     "CP_YZ":
       IF (#compDirection = "LKINCTRL_COMP_LEFT") THEN
         #tempVOrthogonal.x := 0.0;
         #tempVOrthogonal.y := - #tempVTangential.z;
         #tempVOrthogonal.z := #tempVTangential.y;
       ELSE
         #tempVOrthogonal.x := 0.0;
         #tempVOrthogonal.y := #tempVTangential.z;
         #tempVOrthogonal.z := - #tempVTangential.y;
       END_IF;
   END_CASE;
   END_REGION CALCULATION

   #vUnitTangentialPathPlane := #tempVTangential;
   #vUnitOrthogonalPathPlane := #tempVOrthogonal;
   #LKinCtrl_CalcLineTangOrthPathPlane := 0;
END_FUNCTION

FUNCTION "LKinCtrl_CalcCircTangOrthPathPlane" : Word   // FC35056, SCL
TITLE = LKinCtrl_CalcCircTangOrthPathPlane
{ S7_Optimized_Access := 'TRUE' }
AUTHOR : tech.team.motioncontrol@siemens.com
FAMILY : LKinCtrl
VERSION : 1.0
// Calculate orthogonal and tangential vector of a circle point with respect ot the path plane
   VAR_INPUT
      circlePoint : "LKinCtrl_typeCOff3DPoint";   // Circle point
      circleCenterPoint : "LKinCtrl_typeCOff3DPoint";   // Circle center point
      pathPlane : Int;   // Path plane: XZ= 0, YZ=1, XY= 2
      compDirection : Int;   // Tool radius compensation direction: left=1, right = 0
      pathChoice : DInt;   // Circle path choice: positive= 0, negative= 1
   END_VAR
   VAR_OUTPUT
      vUnitTangentialPathPlane : "LKinCtrl_typeCOff3DPoint";   // Output tangential vector - path plane - unit vector
      vUnitOrthogonalPathPlane : "LKinCtrl_typeCOff3DPoint";   // Output othogonal vector - path plane - unit vector
   END_VAR
   VAR_TEMP
      tempDiffVec : "LKinCtrl_typeCOff3DPoint";   // Difference vector
      tempVOrthogonal : "LKinCtrl_typeCOff3DPoint";   // Othogonal vector
      tempVTangential : "LKinCtrl_typeCOff3DPoint";   // Tangential vector
   END_VAR
   // Ret_Val : Return value
   VAR CONSTANT
      ERR_COFF_INVALID_PATH_PLANE : Word := 16#8303;   // Error - invalid path plane
      ERR_COFF_INVALID_PATH_CHOICE_OF_CIRCULAR_CMD : Word := 16#8308;   // Error - invalid circle path choice
      ERR_COFF_INVALID_COMPENSATION_DIRECTION : Word := 16#8304;   // Error - invalid compensation direction
   END_VAR
BEGIN
   //=============================================================================
   // SIEMENS AG
   // (c)Copyright 2019 All Rights Reserved
   //-----------------------------------------------------------------------------
   // Library: - 
   // Tested with: S7-1516T-3 PN
   // Engineering: TIA Portal V15
   // Restrictions: -
   // Requirements: S7-1500/S7-1500T FW 2.5
   // Functionality: Calculate orthogonal and tangential vector of a circle point
   // with respect ot the path plane
   //-----------------------------------------------------------------------------
   // Change log table:
   // Version  Date       Expert in charge Changes applied
   // 01.00.00 2019-02-05 AW               created
   //=============================================================================

   REGION PLAUSIBILITY_CHECK
     // Check path plane
     IF ((#pathPlane >= "CP_XZ") AND (#pathPlane <= "CP_XY"))
     THEN
       // Check compensation direction
       IF ((#compDirection >= "LKINCTRL_COMP_LEFT") AND (#compDirection <= "LKINCTRL_COMP_RIGHT"))
       THEN
         // Check compensation direction
         IF ((#pathChoice >= 0) AND (#pathChoice <= 1))
         THEN
           ;
         ELSE
           #LKinCtrl_CalcCircTangOrthPathPlane := #ERR_COFF_INVALID_PATH_CHOICE_OF_CIRCULAR_CMD; // Invalid compensation direction
           RETURN;
         END_IF;
       ELSE
         #LKinCtrl_CalcCircTangOrthPathPlane := #ERR_COFF_INVALID_COMPENSATION_DIRECTION; // Invalid compensation direction
         RETURN;
       END_IF;
     ELSE
       #LKinCtrl_CalcCircTangOrthPathPlane := #ERR_COFF_INVALID_PATH_PLANE; // Invalid path plane
       RETURN;
     END_IF;
   END_REGION PLAUSIBILITY_CHECK

   REGION CALCULATION



     (*
     IF (#compDirection = "LKINCTRL_COMP_LEFT") THEN
       #tempVOrthogonal := "LKinCtrl_VecSub"(vIn1 := #circlePoint, vIn2 := #circleCenterPoint);
     ELSE
       #tempVOrthogonal := "LKinCtrl_VecSub"(vIn1 := #circleCenterPoint, vIn2 := #circlePoint);
     END_IF;
     *)

     // Take care of path plane
     CASE #pathPlane OF
       "CP_XY":
         // Calc radius vector circle center to start point
         IF (#compDirection = "LKINCTRL_COMP_LEFT") THEN
           IF (#pathChoice = 0) THEN
             #tempVOrthogonal := "LKinCtrl_VecSub"(vIn1 := #circleCenterPoint, vIn2 := #circlePoint);
           ELSE
             #tempVOrthogonal := "LKinCtrl_VecSub"(vIn1 := #circlePoint, vIn2 := #circleCenterPoint);
           END_IF;
         ELSE
           IF (#pathChoice = 0) THEN
             #tempVOrthogonal := "LKinCtrl_VecSub"(vIn1 := #circlePoint, vIn2 := #circleCenterPoint);
           ELSE
             #tempVOrthogonal := "LKinCtrl_VecSub"(vIn1 := #circleCenterPoint, vIn2 := #circlePoint);
           END_IF;
         END_IF;
         #tempVOrthogonal.z := 0.0;

       "CP_XZ":
         // Calc radius vector circle center to start point
         IF (#compDirection = "LKINCTRL_COMP_LEFT") THEN
           IF (#pathChoice = 0) THEN
             #tempVOrthogonal := "LKinCtrl_VecSub"(vIn1 := #circlePoint, vIn2 := #circleCenterPoint);
           ELSE
             #tempVOrthogonal := "LKinCtrl_VecSub"(vIn1 := #circleCenterPoint, vIn2 := #circlePoint);
           END_IF;
         ELSE
           IF (#pathChoice = 0) THEN
             #tempVOrthogonal := "LKinCtrl_VecSub"(vIn1 := #circleCenterPoint, vIn2 := #circlePoint);
           ELSE
             #tempVOrthogonal := "LKinCtrl_VecSub"(vIn1 := #circlePoint, vIn2 := #circleCenterPoint);
           END_IF;
         END_IF;
         #tempVOrthogonal.y := 0.0;

       "CP_YZ":
         // Calc radius vector circle center to start point
         IF (#compDirection = "LKINCTRL_COMP_LEFT") THEN
           IF (#pathChoice = 0) THEN
             #tempVOrthogonal := "LKinCtrl_VecSub"(vIn1 := #circleCenterPoint, vIn2 := #circlePoint);
           ELSE
             #tempVOrthogonal := "LKinCtrl_VecSub"(vIn1 := #circlePoint, vIn2 := #circleCenterPoint);
           END_IF;
         ELSE
           IF (#pathChoice = 0) THEN
             #tempVOrthogonal := "LKinCtrl_VecSub"(vIn1 := #circlePoint, vIn2 := #circleCenterPoint);
           ELSE
             #tempVOrthogonal := "LKinCtrl_VecSub"(vIn1 := #circleCenterPoint, vIn2 := #circlePoint);
           END_IF;
         END_IF;
         #tempVOrthogonal.x := 0.0;
     END_CASE;

     #tempVOrthogonal := "LKinCtrl_VecUnit"(#tempVOrthogonal);

     // Check path plane
     IF (#pathPlane = "CP_XY") THEN
       #tempVTangential.x := - #tempVOrthogonal.y;
       #tempVTangential.y := #tempVOrthogonal.x;
       #tempVTangential.z := 0.0;
     ELSIF (#pathPlane = "CP_XZ") THEN
       #tempVTangential.x := #tempVOrthogonal.z;
       #tempVTangential.y := 0.0;
       #tempVTangential.z := - #tempVOrthogonal.x;
     ELSIF (#pathPlane = "CP_YZ") THEN
       #tempVTangential.x := 0.0;
       #tempVTangential.y := - #tempVOrthogonal.z;
       #tempVTangential.z := #tempVOrthogonal.y;
     END_IF;
   END_REGION CALCULATION

   #vUnitTangentialPathPlane := #tempVTangential;
   #vUnitOrthogonalPathPlane := #tempVOrthogonal;

   #LKinCtrl_CalcCircTangOrthPathPlane := 0; // o.k.
END_FUNCTION

FUNCTION "LKinCtrl_CalcCircCenterByIntermediatePointAndEndPoint" : Word   // FC35057, SCL
TITLE = LKinCtrl_CalcCircCenterByIntermediatePointAndEndPoint
{ S7_Optimized_Access := 'TRUE' }
AUTHOR : tech.team.motioncontrol@siemens.com
FAMILY : LKinCtrl
VERSION : 1.0
// Calculate circle center point with given intermediate point
   VAR_INPUT
      circleStartPoint : "LKinCtrl_typeCOff3DPoint";   // Circle start point
      circleEndPoint : "LKinCtrl_typeCOff3DPoint";   // Circle end point
      circleIntermediatePoint : "LKinCtrl_typeCOff3DPoint";   // Circle intermediate point
      pathPlane : Int;   // Path plane: XZ= 0, YZ=1, XY= 2
   END_VAR
   VAR_OUTPUT
      circleCenterPoint : "LKinCtrl_typeCOff3DPoint";   // Circle center point
   END_VAR
   VAR_TEMP
      tempVecL : "LKinCtrl_typeCOff3DPoint";
      tempVecP1P2 : "LKinCtrl_typeCOff3DPoint";
      tempVecP3P4 : "LKinCtrl_typeCOff3DPoint";
      tempLengthVecP1P2 : LReal;
      tempLengthVecP3P4 : LReal;
      tempUnitVecP1P2 : "LKinCtrl_typeCOff3DPoint";
      tempUnitVecP3P4 : "LKinCtrl_typeCOff3DPoint";
      tempP12 : "LKinCtrl_typeCOff3DPoint";
      tempP34 : "LKinCtrl_typeCOff3DPoint";
      tempP123 : "LKinCtrl_typeCOff3DPoint";
      tempP341 : "LKinCtrl_typeCOff3DPoint";
      tempOrthVecP1P2 : "LKinCtrl_typeCOff3DPoint";
      tempOrthVecP3P4 : "LKinCtrl_typeCOff3DPoint";
      tempRetValue : Word;
      tempPa : "LKinCtrl_typeCOff3DPoint";
      tempPb : "LKinCtrl_typeCOff3DPoint";
      tempMua : LReal;
      tempMub : LReal;
   END_VAR
   // Ret_Val : Return value
   VAR CONSTANT
      ERR_COFF_INVALID_PATH_PLANE : Word := 16#8303;   // Error - invalid path plane
   END_VAR
BEGIN
   //=============================================================================
   // SIEMENS AG
   // (c)Copyright 2019 All Rights Reserved
   //-----------------------------------------------------------------------------
   // Library: - 
   // Tested with: S7-1516T-3 PN
   // Engineering: TIA Portal V15
   // Restrictions: -
   // Requirements: S7-1500/S7-1500T FW 2.5
   // Functionality: Calculate circle center point with given intermediate point
   // and end point
   //-----------------------------------------------------------------------------
   // Change log table:
   // Version  Date       Expert in charge Changes applied
   // 01.00.00 2019-02-05 AW               created
   //=============================================================================


   REGION PLAUSIBILITY_CHECK
   // Check path plane
     IF ((#pathPlane >= "CP_XZ") AND (#pathPlane <= "CP_XY"))
   THEN
     ;
   ELSE
     #LKinCtrl_CalcCircCenterByIntermediatePointAndEndPoint := #ERR_COFF_INVALID_PATH_PLANE; // Invalid path plane
     RETURN;
   END_IF;
   END_REGION PLAUSIBILITY_CHECK

   REGION CALCULATION

     // Intermediate point - start point
     #tempVecP1P2 := "LKinCtrl_VecSub"(vIn1:= #circleIntermediatePoint, vIn2:= #circleStartPoint);
     // Intermediate point - end point
     #tempVecP3P4 := "LKinCtrl_VecSub"(vIn1 := #circleIntermediatePoint, vIn2 := #circleEndPoint);

     // Length of vectors
     #tempLengthVecP1P2 := "LKinCtrl_VecAbs"(#tempVecP1P2);
     #tempLengthVecP3P4 := "LKinCtrl_VecAbs"(#tempVecP3P4);

     // Direction of vectors
     #tempUnitVecP1P2 := "LKinCtrl_VecUnit"(#tempVecP1P2);
     #tempUnitVecP3P4 := "LKinCtrl_VecUnit"(#tempVecP3P4);

     // Perpendicular bisector
     #tempP12 := "LKinCtrl_VecAdd"(vIn1:= #circleStartPoint, vIn2:= "LKinCtrl_VecScale"(vIn:= #tempUnitVecP1P2, factor:= (#tempLengthVecP1P2 / 2.0)));
     #tempP34 := "LKinCtrl_VecAdd"(vIn1:= #circleEndPoint, vIn2:="LKinCtrl_VecScale"(vIn:= #tempUnitVecP3P4, factor:=(#tempLengthVecP3P4 / 2.0)));

     // Rotate vector according to path plane
     // Calc complete shift
     CASE #pathPlane OF
       "CP_XY":
           // Orthogonal end point - intermediate point
           #tempOrthVecP1P2.x := - #tempUnitVecP1P2.y;
           #tempOrthVecP1P2.y := #tempUnitVecP1P2.x;
           #tempOrthVecP1P2.z := 0.0;

           // Orthogonal end point - intermediate point
           #tempOrthVecP3P4.x := #tempUnitVecP3P4.y;
           #tempOrthVecP3P4.y := - #tempUnitVecP3P4.x;
           #tempOrthVecP3P4.z := 0.0;

         "CP_XZ":
           // Orthogonal end point - intermediate point
           #tempOrthVecP1P2.x := #tempUnitVecP1P2.z;
           #tempOrthVecP1P2.y := 0.0;
           #tempOrthVecP1P2.z := - #tempUnitVecP1P2.x;

           // Orthogonal end point - intermediate point
           #tempOrthVecP3P4.x := - #tempUnitVecP3P4.z;
           #tempOrthVecP3P4.y := 0.0;
           #tempOrthVecP3P4.z := #tempUnitVecP3P4.x;

         "CP_YZ":
           // Orthogonal end point - intermediate point
           #tempOrthVecP1P2.x := 0.0;
           #tempOrthVecP1P2.y := - #tempUnitVecP1P2.z;
           #tempOrthVecP1P2.z := #tempUnitVecP1P2.y;

           // Orthogonal end point - intermediate point
           #tempOrthVecP3P4.x := 0.0;
           #tempOrthVecP3P4.y := #tempUnitVecP3P4.z;
           #tempOrthVecP3P4.z := - #tempUnitVecP3P4.y;
     END_CASE;

     #tempOrthVecP1P2 := "LKinCtrl_VecScale"(vIn:= #tempOrthVecP1P2, factor:= #tempLengthVecP1P2);
     #tempOrthVecP3P4 := "LKinCtrl_VecScale"(vIn:= #tempOrthVecP3P4, factor:= #tempLengthVecP3P4);

     #tempP123 := "LKinCtrl_VecAdd"(vIn1:= #tempP12, vIn2:= #tempOrthVecP1P2);
     #tempP341 := "LKinCtrl_VecAdd"(vIn1:= #tempP34, vIn2:= #tempOrthVecP3P4);

     #tempRetValue := "LKinCtrl_CalcLineLineIntersectionPoint"(startPointFirstLine := #tempP12,
                                                      endPointFirstLine := #tempP123,
                                                      startPointSecondLine := #tempP34,
                                                      endPointSecondLine := #tempP341,
                                                      intersectionPointA => #tempPa,
                                                      intersectionPointB => #tempPb,
                                                      muA => #tempMua,
                                                      muB => #tempMub);
     IF (#tempRetValue <> 0) THEN
       #LKinCtrl_CalcCircCenterByIntermediatePointAndEndPoint := #tempRetValue;
       RETURN;
     END_IF;

   END_REGION CALCULATION

   #circleCenterPoint := #tempPa;

   #LKinCtrl_CalcCircCenterByIntermediatePointAndEndPoint := 0; // o.k.
END_FUNCTION

FUNCTION "LKinCtrl_CalcCircPathChoiceByIntermediatePointAndEndPoint" : Word   // FC35058, SCL
TITLE = LKinCtrl_CalcCircPathChoiceByIntermediatePointAndEndPoint
{ S7_Optimized_Access := 'TRUE' }
AUTHOR : tech.team.motioncontrol@siemens.com
FAMILY : LKinCtrl
VERSION : 1.0
// Calculate circle path choice by given circle intermediate point and end point
   VAR_INPUT
      circleStartPoint : "LKinCtrl_typeCOff3DPoint";   // Circle start point
      circleEndPoint : "LKinCtrl_typeCOff3DPoint";   // Circle end point
      circleintermediatePoint : "LKinCtrl_typeCOff3DPoint";   // Circle intermediate point
      pathPlane : Int;   // Path plane: XZ= 0, YZ=1, XY= 2
   END_VAR
   VAR_OUTPUT
      pathChoice : DInt;   // Circle path choice: positive= 0, negative= 1
   END_VAR
   VAR_TEMP
      tempVEndStart : "LKinCtrl_typeCOff3DPoint";
      tempVIntStart : "LKinCtrl_typeCOff3DPoint";
      tempCrossVec : "LKinCtrl_typeCOff3DPoint";
   END_VAR
   // Ret_Val : Return value
   VAR CONSTANT
      ERR_COFF_INVALID_PATH_PLANE : Word := 16#8303;   // Error - invalid path plane
   END_VAR
BEGIN
   //=============================================================================
   // SIEMENS AG
   // (c)Copyright 2019 All Rights Reserved
   //-----------------------------------------------------------------------------
   // Library: - 
   // Tested with: S7-1516T-3 PN
   // Engineering: TIA Portal V15
   // Restrictions: -
   // Requirements: S7-1500/S7-1500T FW 2.5
   // Functionality: Calculate circle path choice by given circle intermediate point
   // and end point
   //-----------------------------------------------------------------------------
   // Change log table:
   // Version  Date       Expert in charge Changes applied
   // 01.00.00 2019-02-05 AW               created
   //=============================================================================

   REGION PLAUSIBILITY_CHECK
     // Check path plane
     IF ((#pathPlane >= "CP_XZ") AND (#pathPlane <= "CP_XY"))
     THEN
       ;
     ELSE
       #LKinCtrl_CalcCircPathChoiceByIntermediatePointAndEndPoint := #ERR_COFF_INVALID_PATH_PLANE; // Invalid path plane
       RETURN;
     END_IF;
   END_REGION PLAUSIBILITY_CHECK

   REGION CALCULATION

   (*  
   // Calculate angle between start / end point and start / intermediate point
     #tempRetValue := "LKinCOff_CalcAngleBetweenVectors"(point1 := #endPoint,
                                                         point2 := #intermediatePoint,
                                                         intersectionPoint := #startPoint,
                                                         angle => #tempAngle);


   IF (#tempRetValue <> 0) THEN
     #LKinCOff_CalcPathChoiceByIntermediatePointAndEndPoint := #tempRetValue;
     RETURN;
   END_IF;

   END_REGION CALCULATION
   IF (#tempAngle < 0.0) THEN
     #pathChoice := 1;
   ELSE
     #pathChoice := 0;
   END_IF;
   *)

     // Difference vectors
     #tempVEndStart := "LKinCtrl_VecSub"(vIn1 := #circleEndPoint, vIn2 := #circleStartPoint);
     #tempVIntStart := "LKinCtrl_VecSub"(vIn1 := #circleintermediatePoint, vIn2 := #circleStartPoint);

     #tempCrossVec := "LKinCtrl_VecCrossProd"(vIn1 := #tempVEndStart,
                                              vIn2 := #tempVIntStart);

     // Check path plane
     IF (#pathPlane = "CP_XY") THEN
       IF (#tempCrossVec.z > 0.0) THEN
         #pathChoice := "PC_NEGATIVE";
       ELSE
         #pathChoice := "PC_POSITIVE";
       END_IF;
     ELSIF (#pathPlane = "CP_XZ") THEN
       IF (#tempCrossVec.y > 0.0) THEN
         #pathChoice := "PC_NEGATIVE";
       ELSE
         #pathChoice := "PC_POSITIVE";
       END_IF;
     ELSIF (#pathPlane = "CP_YZ") THEN
       IF (#tempCrossVec.x > 0.0) THEN
         #pathChoice := "PC_NEGATIVE";
       ELSE
         #pathChoice := "PC_POSITIVE";
       END_IF;
     END_IF;

    END_REGION; 
   #LKinCtrl_CalcCircPathChoiceByIntermediatePointAndEndPoint := 0; // o.k.
END_FUNCTION

FUNCTION "LKinCtrl_CalcAngleBetweenVectors" : Word   // FC35059, SCL
TITLE = LKinCtrl_CalcAngleBetweenVectors
{ S7_Optimized_Access := 'TRUE' }
AUTHOR : tech.team.motioncontrol@siemens.com
FAMILY : LKinCtrl
VERSION : 1.0
// Calculate angle between two intersecting vectors
   VAR_INPUT
      point1 : "LKinCtrl_typeCOff3DPoint";   // Point 1
      point2 : "LKinCtrl_typeCOff3DPoint";   // Point 2
      intersectionPoint : "LKinCtrl_typeCOff3DPoint";   // Common point
   END_VAR
   VAR_OUTPUT
      angle : LReal;   // Calculated angle
   END_VAR
   VAR_TEMP
      tempVecP1InterPoint : "LKinCtrl_typeCOff3DPoint";
      tempVecP2InterPoint : "LKinCtrl_typeCOff3DPoint";
      tempValue : LReal;
      tempVecP1P2 : "LKinCtrl_typeCOff3DPoint";
      tempVecP3P4 : "LKinCtrl_typeCOff3DPoint";
      tempLengthVecP1P2 : LReal;
      tempLengthVecP3P4 : LReal;
      tempUnitVecP1P2 : "LKinCtrl_typeCOff3DPoint";
      tempUnitVecP3P4 : "LKinCtrl_typeCOff3DPoint";
      tempP12 : "LKinCtrl_typeCOff3DPoint";
      tempP34 : "LKinCtrl_typeCOff3DPoint";
      tempP123 : "LKinCtrl_typeCOff3DPoint";
      tempP341 : "LKinCtrl_typeCOff3DPoint";
      tempOrthVecP1P2 : "LKinCtrl_typeCOff3DPoint";
      tempOrthVecP3P4 : "LKinCtrl_typeCOff3DPoint";
      tempRetValue : Int;
      tempPa1 : "LKinCtrl_typeCOff3DPoint";
      tempPb1 : "LKinCtrl_typeCOff3DPoint";
      tempMua : LReal;
      TempMub : LReal;
   END_VAR
   // Ret_Val : Return value
   VAR CONSTANT
      ERR_COFF_VECTOR_LENGTH_ZERO : Word := 16#8310;   // Error - vector length is zero
      ERR_COFF_INVALID_ACOS_ARGUMENT : Word := 16#8311;   // Error - invalid ACOS argument
   END_VAR
BEGIN
   //=============================================================================
   // SIEMENS AG
   // (c)Copyright 2019 All Rights Reserved
   //-----------------------------------------------------------------------------
   // Library: - 
   // Tested with: S7-1516T-3 PN
   // Engineering: TIA Portal V15
   // Restrictions: -
   // Requirements: S7-1500/S7-1500T FW 2.5
   // Functionality: Calculate angle between two intersecting vectors
   //-----------------------------------------------------------------------------
   // Change log table:
   // Version  Date       Expert in charge Changes applied
   // 01.00.00 2019-02-05 AW               created
   //=============================================================================
   REGION PLAUSIBILITY_CHECK
   END_REGION PLAUSIBILITY_CHECK

   REGION CALCULATION

     // Difference vectors
     // Point 1 - intersection point
     #tempVecP1InterPoint := "LKinCtrl_VecSub"(vIn1:= #point1, vIn2:= #intersectionPoint);
     // Point 2 - intersection point
     #tempVecP2InterPoint := "LKinCtrl_VecSub"(vIn1 := #point2, vIn2 := #intersectionPoint);

     #tempValue := "LKinCtrl_VecAbs"(#tempVecP1InterPoint) * "LKinCtrl_VecAbs"(#tempVecP2InterPoint);

     IF (#tempValue = 0.0) THEN
       #LKinCtrl_CalcAngleBetweenVectors := #ERR_COFF_VECTOR_LENGTH_ZERO; // division by zero
       RETURN;
     END_IF;

     #tempValue := "LKinCtrl_VecScalProd"(vIn1:=#tempVecP1InterPoint, vIn2:=#tempVecP2InterPoint) / #tempValue;

     IF ((#tempValue < -1.0) OR (#tempValue > 1.0)) THEN
       #LKinCtrl_CalcAngleBetweenVectors := #ERR_COFF_INVALID_ACOS_ARGUMENT; // acos only defined for -1 ... +1
       RETURN;
     ELSE
       // Angle between vector 1 and vector 2
       #angle := ACOS(#tempValue) * 180.0 / "LKINCTRL_PI";
     END_IF;

   END_REGION CALCULATION



   #LKinCtrl_CalcAngleBetweenVectors := 0; // o.k.
END_FUNCTION

FUNCTION "LKinCtrl_CalcLineLineIntersectionPoint" : Word   // FC35060, SCL
TITLE = LKinCtrl_CalcLineLineIntersectionPoint
{ S7_Optimized_Access := 'TRUE' }
AUTHOR : tech.team.motioncontrol@siemens.com
FAMILY : LKinCtrl
VERSION : 1.0
// Calculate the line segment Pa/Pb that is the shortest route between two lines P1P2 and P3P4
   VAR_INPUT
      startPointFirstLine : "LKinCtrl_typeCOff3DPoint";   // Start point first line
      endPointFirstLine : "LKinCtrl_typeCOff3DPoint";   // End point first line
      startPointSecondLine : "LKinCtrl_typeCOff3DPoint";   // Start point second line
      endPointSecondLine : "LKinCtrl_typeCOff3DPoint";   // End point second line
   END_VAR
   VAR_OUTPUT
      intersectionPointA : "LKinCtrl_typeCOff3DPoint";   // Intersection point a
      intersectionPointB : "LKinCtrl_typeCOff3DPoint";   // Intersection point b
      muA : LReal;   // Direction vector a
      muB : LReal;   // Direction vector b
   END_VAR
   VAR_TEMP
      tempP13 : "LKinCtrl_typeCOff3DPoint";
      tempP43 : "LKinCtrl_typeCOff3DPoint";
      tempP21 : "LKinCtrl_typeCOff3DPoint";
      tempD1343 : LReal;
      tempD4321 : LReal;
      tempD1321 : LReal;
      tempD4343 : LReal;
      tempD2121 : LReal;
      tempNumer : LReal;
      tempDenom : LReal;
   END_VAR
   // Ret_Val : Return value
   VAR CONSTANT
      COFF_EPS : LReal := 0.001;   // Internal constant
      ERR_COFF_LINES_DO_NOT_INTERSECT : Word := 16#8312;   // Error - no solution, lines don't intersect
      ERR_COFF_ZERO_VECTOR : Word := 16#8313;   // Error - zero vector
   END_VAR
BEGIN
   //=============================================================================
   // SIEMENS AG
   // (c)Copyright 2019 All Rights Reserved
   //-----------------------------------------------------------------------------
   // Library: - 
   // Tested with: S7-1516T-3 PN
   // Engineering: TIA Portal V15
   // Restrictions: -
   // Requirements: S7-1500/S7-1500T FW 2.5
   // Functionality: Calculate the line segment Pa/Pb that is the shortest route
   // between two lines P1P2 and P3P4. Calculate also the values of mua and mub where
   // Pa = P1 + mua (P2 - P1)
   // Pb = P3 + mub (P4 - P3)
   // Return error if the lines don't intersect
   //-----------------------------------------------------------------------------
   // Change log table:
   // Version  Date       Expert in charge Changes applied
   // 01.00.00 2019-02-05 AW               created
   //=============================================================================
   REGION PLAUSIBILITY_CHECK

   END_REGION PLAUSIBILITY_CHECK

   REGION CALCULATION
     #tempP13.x := #startPointFirstLine.x - #startPointSecondLine.x;
     #tempP13.y := #startPointFirstLine.y - #startPointSecondLine.y;
     #tempP13.z := #startPointFirstLine.z - #startPointSecondLine.z;
     #tempP43.x := #endPointSecondLine.x - #startPointSecondLine.x;
     #tempP43.y := #endPointSecondLine.y - #startPointSecondLine.y;
     #tempP43.z := #endPointSecondLine.z - #startPointSecondLine.z;
     IF ((ABS(#tempP43.x) < #COFF_EPS) AND (ABS(#tempP43.y) < #COFF_EPS) AND (ABS(#tempP43.z) < #COFF_EPS)) THEN
       #LKinCtrl_CalcLineLineIntersectionPoint := #ERR_COFF_LINES_DO_NOT_INTERSECT;
       RETURN;
     END_IF;

     #tempP21.x := #endPointFirstLine.x - #startPointFirstLine.x;
     #tempP21.y := #endPointFirstLine.y - #startPointFirstLine.y;
     #tempP21.z := #endPointFirstLine.z - #startPointFirstLine.z;
     IF ((ABS(#tempP21.x) < #COFF_EPS) AND (ABS(#tempP21.y) < #COFF_EPS) AND (ABS(#tempP21.z) < #COFF_EPS)) THEN
       #LKinCtrl_CalcLineLineIntersectionPoint := #ERR_COFF_LINES_DO_NOT_INTERSECT;
       RETURN;
     END_IF;

     #tempD1343 := #tempP13.x * #tempP43.x + #tempP13.y * #tempP43.y + #tempP13.z * #tempP43.z;
     #tempD4321 := #tempP43.x * #tempP21.x + #tempP43.y * #tempP21.y + #tempP43.z * #tempP21.z;
     #tempD1321 := #tempP13.x * #tempP21.x + #tempP13.y * #tempP21.y + #tempP13.z * #tempP21.z;
     #tempD4343 := #tempP43.x * #tempP43.x + #tempP43.y * #tempP43.y + #tempP43.z * #tempP43.z;
     #tempD2121 := #tempP21.x * #tempP21.x + #tempP21.y * #tempP21.y + #tempP21.z * #tempP21.z;

     #tempDenom := #tempD2121 * #tempD4343 - #tempD4321 * #tempD4321;
     IF (ABS(#tempDenom) < #COFF_EPS) THEN
       #LKinCtrl_CalcLineLineIntersectionPoint := #ERR_COFF_LINES_DO_NOT_INTERSECT;
       RETURN;
     END_IF;

     #tempNumer := #tempD1343 * #tempD4321 - #tempD1321 * #tempD4343;

     #muA := #tempNumer / #tempDenom;
     #muB := (#tempD1343 + #tempD4321 * #muA) / #tempD4343;

     #intersectionPointA.x := #startPointFirstLine.x + #muA * #tempP21.x;
     #intersectionPointA.y := #startPointFirstLine.y + #muA * #tempP21.y;
     #intersectionPointA.z := #startPointFirstLine.z + #muA * #tempP21.z;

     #intersectionPointB.x := #startPointSecondLine.x + #muB * #tempP43.x;
     #intersectionPointB.y := #startPointSecondLine.y + #muB * #tempP43.y;
     #intersectionPointB.z := #startPointSecondLine.z + #muB * #tempP43.z;

   END_REGION
   #LKinCtrl_CalcLineLineIntersectionPoint := 0;
END_FUNCTION

FUNCTION "LKinCtrl_CalcLineCircleIntersectionPoint" : Word   // FC35061, SCL
TITLE = LKinCtrl_CalcLineCircleIntersectionPoint
{ S7_Optimized_Access := 'TRUE' }
AUTHOR : tech.team.motioncontrol@siemens.com
FAMILY : LKinCtrl
VERSION : 1.1
// Calculate the intersection of a ray and a sphere
   VAR_INPUT
      startPointLine : "LKinCtrl_typeCOff3DPoint";   // Start point line
      endPointLine : "LKinCtrl_typeCOff3DPoint";   // End point line
      circleCenter : "LKinCtrl_typeCOff3DPoint";   // Circle center
      circleRadius : LReal;   // Circle radius
   END_VAR
   VAR_OUTPUT
      intersectionPointA : "LKinCtrl_typeCOff3DPoint";   // Intersection point a
      intersectionPointB : "LKinCtrl_typeCOff3DPoint";   // Intersection point b
   END_VAR
   VAR_TEMP
      tempP13 : "LKinCtrl_typeCOff3DPoint";
      tempP43 : "LKinCtrl_typeCOff3DPoint";
      tempA : LReal;
      tempB : LReal;
      tempC : LReal;
      tempBb4ac : LReal;
      tempDp : "LKinCtrl_typeCOff3DPoint";
      tempP22 : "LKinCtrl_typeCOff3DPoint";
      tempMuA : LReal;
      tempMuB : LReal;
   END_VAR
   // Ret_Val : Return value
   VAR CONSTANT
      COFF_EPS : LReal := 0.001;   // Internal constant
      ERR_COFF_LINE_CIRCLE_DO_NOT_INTERSECT : Word := 16#8315;   // Error - no solution - line and circle don't intersect
   END_VAR
BEGIN
   //=============================================================================
   // SIEMENS AG
   // (c)Copyright 2019 All Rights Reserved
   //-----------------------------------------------------------------------------
   // Library: - 
   // Tested with: S7-1516T-3 PN
   // Engineering: TIA Portal V15
   // Restrictions: -
   // Requirements: S7-1500/S7-1500T FW 2.5
   // Functionality: Calculate the intersection of a ray and a sphere
   // The line segment is defined from p1 to p2
   // The sphere is of radius r and centered at sc
   // There are potentially two points of intersection given by
   // p = p1 + mu1 (p2 - p1)
   // p = p1 + mu2 (p2 - p1)
   // Return error if the ray doesn't intersect the sphere.
   //-----------------------------------------------------------------------------
   // Change log table:
   // Version  Date       Expert in charge Changes applied
   // 01.00.00 2019-02-05 AW               created
   // 01.01.00 2020-07-24 AW               #tempBb4ac fix (<= --> <) and tolerance added
   //=============================================================================

   REGION CALCULATION  
     #tempDp.x := #endPointLine.x - #startPointLine.x;
     #tempDp.y := #endPointLine.y - #startPointLine.y;
     #tempDp.z := #endPointLine.z - #startPointLine.z;
     #tempA := #tempDp.x * #tempDp.x + #tempDp.y * #tempDp.y + #tempDp.z * #tempDp.z;


     #tempB := 2.0 * (#tempDp.x * (#startPointLine.x - #circleCenter.x) + #tempDp.y * (#startPointLine.y - #circleCenter.y) + #tempDp.z * (#startPointLine.z - #circleCenter.z));
     #tempC := #circleCenter.x * #circleCenter.x + #circleCenter.y * #circleCenter.y + #circleCenter.z * #circleCenter.z;
     #tempC := #tempC + #startPointLine.x * #startPointLine.x + #startPointLine.y * #startPointLine.y + #startPointLine.z * #startPointLine.z;
     #tempC := #tempC - 2.0 * (#circleCenter.x * #startPointLine.x + #circleCenter.y * #startPointLine.y + #circleCenter.z * #startPointLine.z);
     #tempC := #tempC - #circleRadius * #circleRadius;
     #tempBb4ac := #tempB * #tempB - 4.0 * #tempA * #tempC;

     IF ((ABS(#tempA) < #COFF_EPS))
     THEN
       #tempMuA := 0;
       #tempMuB := 0;
       #LKinCtrl_CalcLineCircleIntersectionPoint := #ERR_COFF_LINE_CIRCLE_DO_NOT_INTERSECT;
       RETURN;
     END_IF;

     // Three possible solution:
     // #tempBb4ac > 0 - two intersection points
     // #tempBb4ax = 0 - one intersection point (additional tolerance)
     // #tempBb4ax < 0 - no intersection point (additional tolerance) 

     // 01.00.01 2020-07-24
     IF (#tempBb4ac < 0.0) THEN
       // Within tolerance (accept tiny floating point deviations)
       IF (ABS(#tempBb4ac) < #COFF_EPS) THEN
         #tempBb4ac := 0.0;
       ELSE
         #LKinCtrl_CalcLineCircleIntersectionPoint := #ERR_COFF_LINE_CIRCLE_DO_NOT_INTERSECT;
         RETURN;
       END_IF;
     END_IF;


     #tempMuA := (- #tempB + SQRT(#tempBb4ac)) / (2.0 * #tempA);
     #tempMuB := (- #tempB - SQRT(#tempBb4ac)) / (2.0 * #tempA);
     //pa  := p1 + mu1 (p2 - p1)
     //pb  := p1 + mu2 (p2 - p1)


     #intersectionPointA.x := #startPointLine.x + #tempMuA * #tempDp.x;
     #intersectionPointA.y := #startPointLine.y + #tempMuA * #tempDp.y;
     #intersectionPointA.z := #startPointLine.z + #tempMuA * #tempDp.z;
     #intersectionPointB.x := #startPointLine.x + #tempMuB * #tempDp.x;
     #intersectionPointB.y := #startPointLine.y + #tempMuB * #tempDp.y;
     #intersectionPointB.z := #startPointLine.z + #tempMuB * #tempDp.z;

   END_REGION

   #LKinCtrl_CalcLineCircleIntersectionPoint := 0;
END_FUNCTION

FUNCTION "LKinCtrl_CalcCircleCircleIntersectionPoint" : Word   // FC35062, SCL
TITLE = LKinCtrl_CalcCircleCircleIntersectionPoint
{ S7_Optimized_Access := 'TRUE' }
AUTHOR : tech.team.motioncontrol@siemens.com
FAMILY : LKinCtrl
VERSION : 1.1
// Determine the points where 2 circles in a common plane intersect
   VAR_INPUT
      circleCenterPoint1 : "LKinCtrl_typeCOff3DPoint";   // Center point of first circle
      circleCenterPoint2 : "LKinCtrl_typeCOff3DPoint";   // Center point of second circle
      circleRadius1 : LReal;   // Radius of first circle
      circleRadius2 : LReal;   // Radius of second circle
      pathPlane : Int;   // Path plane: XZ= 0, YZ=1, XY= 2
   END_VAR
   VAR_OUTPUT
      intersectionPointA : "LKinCtrl_typeCOff3DPoint";   // Intersection point a
      intersectionPointB : "LKinCtrl_typeCOff3DPoint";   // Intersection point b
   END_VAR
   VAR_TEMP
      tempP02 : LReal;
      tempvDiff : "LKinCtrl_typeCOff3DPoint";
      tempCenterDistance : LReal;
      tempH : LReal;
      tempInterPointOffset : "LKinCtrl_typeCOff3DPoint";
      tempP2 : "LKinCtrl_typeCOff3DPoint";
   END_VAR
   // Ret_Val : Return value
   VAR CONSTANT
      COFF_EPS : LReal := 0.001;   // Internal constant
      ERR_COFF_INVALID_PATH_PLANE : Word := 16#8303;   // Error - invalid path plane
      ERR_COFF_CIRCLES_DO_NOT_INTERSECT : Word := 16#8318;   // Error - no solution - circles don't intersect
      ERR_COFF_ONE_CIRC_CONTAINED_IN_THE_OTHER : Word := 16#8319;   // Error - one circle is contained in the other
      ERR_COFF_CIRCLE_CENTERS_EQUAL : Word := 16#8350;   // Error - circle centers are equal infinite intersections (only internal)
   END_VAR
BEGIN
   //=============================================================================
   // SIEMENS AG
   // (c)Copyright 2019 All Rights Reserved
   //-----------------------------------------------------------------------------
   // Library: - 
   // Tested with: S7-1516T-3 PN
   // Engineering: TIA Portal V15
   // Restrictions: -
   // Requirements: S7-1500/S7-1500T FW 2.5
   // Functionality: Determine the points where 2 circles in a common plane intersect
   // center and radius of 1st circle
   // center and radius of 2nd circle
   // 1st intersection point - pa
   // 2nd intersection point - pb
   //-----------------------------------------------------------------------------
   // Change log table:
   // Version  Date       Expert in charge Changes applied
   // 01.00.00 2019-02-05 AW               created
   // 01.01.00 2020-08-14 AW               bugfix equal circle centers
   // 01.01.01 2020-08-25 AW               bugfix tiny floating point deviations due to calculation - circles intersect in one point
   //=============================================================================

   REGION PLAUSIBILITY_CHECK
     // Check path plane
     IF ((#pathPlane >= "CP_XZ") AND (#pathPlane <= "CP_XY"))
     THEN
       ;
     ELSE
       #LKinCtrl_CalcCircleCircleIntersectionPoint := #ERR_COFF_INVALID_PATH_PLANE; // Invalid path plane
       RETURN;
     END_IF;
   END_REGION PLAUSIBILITY_CHECK

   REGION CALCULATION   
     // Distinguish between different path planes
     CASE #pathPlane OF
       "CP_XY":
         // dx and dy are the vertical and horizontal distances between the circle centers
         #tempvDiff.x := #circleCenterPoint2.x - #circleCenterPoint1.x;
         #tempvDiff.y := #circleCenterPoint2.y - #circleCenterPoint1.y;

         // Determine the straight-line distance between the centers.
         #tempCenterDistance := SQRT((#tempvDiff.y * #tempvDiff.y) + (#tempvDiff.x * #tempvDiff.x));

         // No solution possible - circles do not intersect
         IF (#tempCenterDistance > (#circleRadius1 + #circleRadius2)) THEN
           // V01.01.01
           IF (#tempCenterDistance < (#circleRadius1 + #circleRadius2 + #COFF_EPS)) THEN
             #tempCenterDistance := #circleRadius1 + #circleRadius2;
           ELSE
             #LKinCtrl_CalcCircleCircleIntersectionPoint := #ERR_COFF_CIRCLES_DO_NOT_INTERSECT;
             RETURN;
           END_IF;
         END_IF;

         // No solution - one circle is contained in the other
         IF (#tempCenterDistance < ABS(#circleRadius1 - #circleRadius2)) THEN
           // V01.01.01
           IF (#tempCenterDistance > (ABS(#circleRadius1 - #circleRadius2) - #COFF_EPS)) THEN
             #tempCenterDistance := ABS(#circleRadius1 - #circleRadius2);
           ELSE
             #LKinCtrl_CalcCircleCircleIntersectionPoint := #ERR_COFF_ONE_CIRC_CONTAINED_IN_THE_OTHER;
             RETURN;
           END_IF;
         END_IF;

         // Both circle centers are equal
         IF (#tempCenterDistance <= 0.0) THEN
           #LKinCtrl_CalcCircleCircleIntersectionPoint := #ERR_COFF_CIRCLE_CENTERS_EQUAL;
           RETURN;
         END_IF;

         // 'point 2' is the point where the line through the circle
         // intersection points crosses the line between the circle centers.  

         // Determine the distance from point 0 to point 2
         #tempP02 := ((#circleRadius1 * #circleRadius1) - (#circleRadius2 * #circleRadius2) + (#tempCenterDistance * #tempCenterDistance)) / (2.0 * #tempCenterDistance);

         // Determine the coordinates of point 2
         #tempP2.x := #circleCenterPoint1.x + (#tempvDiff.x * #tempP02 / #tempCenterDistance);
         #tempP2.y := #circleCenterPoint1.y + (#tempvDiff.y * #tempP02 / #tempCenterDistance);

         // Determine the distance from point 2 to either of the intersection points
         #tempH := SQRT((#circleRadius1 * #circleRadius1) - (#tempP02 * #tempP02));

         // Determine the offsets of the intersection points from point 2
         #tempInterPointOffset.x := - #tempvDiff.y * (#tempH / #tempCenterDistance);
         #tempInterPointOffset.y := #tempvDiff.x * (#tempH / #tempCenterDistance);

         // Determine the absolute intersection points
         #intersectionPointA.x := #tempP2.x + #tempInterPointOffset.x;
         #intersectionPointB.x := #tempP2.x - #tempInterPointOffset.x;
         #intersectionPointA.y := #tempP2.y + #tempInterPointOffset.y;
         #intersectionPointB.y := #tempP2.y - #tempInterPointOffset.y;

           // Get third coordinate
           #intersectionPointA.z := #circleCenterPoint1.z;
           #intersectionPointB.z := #circleCenterPoint1.z;

       "CP_XZ":
         // dz AND dx are the vertical and horizontal distances between the circle centers
         #tempvDiff.z := #circleCenterPoint2.z - #circleCenterPoint1.z;
         #tempvDiff.x := #circleCenterPoint2.x - #circleCenterPoint1.x;

         // Determine the straight-line distance between the centers.
         #tempCenterDistance := SQRT((#tempvDiff.x * #tempvDiff.x) + (#tempvDiff.z * #tempvDiff.z));

         // No solution possible - circles do not intersect
         IF (#tempCenterDistance > (#circleRadius1 + #circleRadius2)) THEN
           // V01.01.01
           IF (#tempCenterDistance < (#circleRadius1 + #circleRadius2 + #COFF_EPS)) THEN
             #tempCenterDistance := #circleRadius1 + #circleRadius2;
           ELSE
             #LKinCtrl_CalcCircleCircleIntersectionPoint := #ERR_COFF_CIRCLES_DO_NOT_INTERSECT;
             RETURN;
           END_IF;
         END_IF;

         // No solution - one circle is contained in the other
         IF (#tempCenterDistance < ABS(#circleRadius1 - #circleRadius2)) THEN
           // V01.01.01
           IF (#tempCenterDistance > (ABS(#circleRadius1 - #circleRadius2) - #COFF_EPS)) THEN
             #tempCenterDistance := ABS(#circleRadius1 - #circleRadius2);
           ELSE
             #LKinCtrl_CalcCircleCircleIntersectionPoint := #ERR_COFF_ONE_CIRC_CONTAINED_IN_THE_OTHER;
             RETURN;
           END_IF;
         END_IF;

         // Both circle centers are equal
         IF (#tempCenterDistance <= 0.0) THEN
           #LKinCtrl_CalcCircleCircleIntersectionPoint := #ERR_COFF_CIRCLE_CENTERS_EQUAL;
           RETURN;
         END_IF;

         // 'point 2' is the point where the line through the circle
         // intersection points crosses the line between the circle centers.  

         // Determine the distance from point 0 to point 2
         #tempP02 := ((#circleRadius1 * #circleRadius1) - (#circleRadius2 * #circleRadius2) + (#tempCenterDistance * #tempCenterDistance)) / (2.0 * #tempCenterDistance);

         // Determine the coordinates of point 2
         #tempP2.z := #circleCenterPoint1.z + (#tempvDiff.z * #tempP02 / #tempCenterDistance);
         #tempP2.x := #circleCenterPoint1.x + (#tempvDiff.x * #tempP02 / #tempCenterDistance);

         // Determine the distance from point 2 to either of the intersection points
         #tempH := SQRT((#circleRadius1 * #circleRadius1) - (#tempP02 * #tempP02));

         // Determine the offsets of the intersection points from point 2
         // Before
         #tempInterPointOffset.z := - #tempvDiff.x * (#tempH / #tempCenterDistance);
         #tempInterPointOffset.x := #tempvDiff.z * (#tempH / #tempCenterDistance);

         // Determine the absolute intersection points
         #intersectionPointA.z := #tempP2.z + #tempInterPointOffset.z;
         #intersectionPointB.z := #tempP2.z - #tempInterPointOffset.z;
         #intersectionPointA.x := #tempP2.x + #tempInterPointOffset.x;
         #intersectionPointB.x := #tempP2.x - #tempInterPointOffset.x;

         // Get third coordinate
         #intersectionPointA.y := #circleCenterPoint1.y;
         #intersectionPointB.y := #circleCenterPoint1.y;

       "CP_YZ":
         // dx AND dy are the vertical and horizontal distances between the circle centers
         #tempvDiff.y := #circleCenterPoint2.y - #circleCenterPoint1.y;
         #tempvDiff.z := #circleCenterPoint2.z - #circleCenterPoint1.z;

         // Determine the straight-line distance between the centers.
         #tempCenterDistance := SQRT((#tempvDiff.z * #tempvDiff.z) + (#tempvDiff.y * #tempvDiff.y));

         // No solution possible - circles do not intersect
         IF (#tempCenterDistance > (#circleRadius1 + #circleRadius2)) THEN
           // V01.01.01
           IF (#tempCenterDistance < (#circleRadius1 + #circleRadius2 + #COFF_EPS)) THEN
             #tempCenterDistance := #circleRadius1 + #circleRadius2;
           ELSE
             #LKinCtrl_CalcCircleCircleIntersectionPoint := #ERR_COFF_CIRCLES_DO_NOT_INTERSECT;
             RETURN;
           END_IF;
         END_IF;

         // No solution - one circle is contained in the other
         IF (#tempCenterDistance < ABS(#circleRadius1 - #circleRadius2)) THEN
           // V01.01.01
           IF (#tempCenterDistance > (ABS(#circleRadius1 - #circleRadius2) - #COFF_EPS)) THEN
             #tempCenterDistance := ABS(#circleRadius1 - #circleRadius2);
           ELSE
             #LKinCtrl_CalcCircleCircleIntersectionPoint := #ERR_COFF_ONE_CIRC_CONTAINED_IN_THE_OTHER;
             RETURN;
           END_IF;
         END_IF;

         // Both circle centers are equal
         IF (#tempCenterDistance <= 0.0) THEN
           #LKinCtrl_CalcCircleCircleIntersectionPoint := #ERR_COFF_CIRCLE_CENTERS_EQUAL;
           RETURN;
         END_IF;

         // 'point 2' is the point where the line through the circle
         // intersection points crosses the line between the circle centers.  

         // Determine the distance from point 0 to point 2
         #tempP02 := ((#circleRadius1 * #circleRadius1) - (#circleRadius2 * #circleRadius2) + (#tempCenterDistance * #tempCenterDistance)) / (2.0 * #tempCenterDistance);

         // Determine the coordinates of point 2
         #tempP2.y := #circleCenterPoint1.y + (#tempvDiff.y * #tempP02 / #tempCenterDistance);
         #tempP2.z := #circleCenterPoint1.z + (#tempvDiff.z * #tempP02 / #tempCenterDistance);

         // Determine the distance from point 2 to either of the intersection points
         #tempH := SQRT((#circleRadius1 * #circleRadius1) - (#tempP02 * #tempP02));

         // Determine the offsets of the intersection points from point 2
         #tempInterPointOffset.y := - #tempvDiff.z * (#tempH / #tempCenterDistance);
         #tempInterPointOffset.z := #tempvDiff.y * (#tempH / #tempCenterDistance);

         // Determine the absolute intersection points
         #intersectionPointA.y := #tempP2.y + #tempInterPointOffset.y;
         #intersectionPointB.y := #tempP2.y - #tempInterPointOffset.y;
         #intersectionPointA.z := #tempP2.z + #tempInterPointOffset.z;
         #intersectionPointB.z := #tempP2.z - #tempInterPointOffset.z;

         // Get third coordinate
         #intersectionPointA.x := #circleCenterPoint1.x;
         #intersectionPointB.x := #circleCenterPoint1.x;
     END_CASE;
   END_REGION

   #LKinCtrl_CalcCircleCircleIntersectionPoint := 16#0;
END_FUNCTION

FUNCTION "LKinCtrl_CartesianCoordTo3DPoint" : "LKinCtrl_typeCOff3DPoint"   // FC35065, SCL
TITLE = LKinCtrl_CartesianCoordTo3DPoint
{ S7_Optimized_Access := 'TRUE' }
AUTHOR : tech.team.motioncontrol@siemens.com
FAMILY : LKinCtrl
VERSION : 1.0
// The function converts data type "LKinCtrl_typeCartesianPosition" in "LKinCtrl_typeCOff3DPoint"
   VAR_INPUT
      cartesianCoord : "LKinCtrl_typeCartesianPosition";   // Cartesian input coordinate
   END_VAR
   // Ret_Val : Return - 3D output point
BEGIN
   //==========================================================================================
   // SIEMENS AG
   // (c)Copyright 2019 All Rights Reserved
   //------------------------------------------------------------------------------------------
   // Library: LCOffset
   // Tested with: S7-1515T-3 PN/DP
   // Engineering: TIA Portal V15
   // Restrictions: ---
   // Requirements: S7-1500T FW 2.5
   // Functionality: The function converts data type "LKinCtrl_typeCartesianPosition" in "LKinCtrl_typeCOff3DPoint"
   // Support: tech.team.motioncontrol@siemens.com
   // Note: Parameter comments are only available in language 'English (United States)'
   //------------------------------------------------------------------------------------------
   // Change log table:
   // Version    Date          Expert in charge    Changes applied
   // 01.00.00   2019-02-14    AW                  created
   //===========================================================================================
   //
   #LKinCtrl_CartesianCoordTo3DPoint.x := #cartesianCoord.x;
   #LKinCtrl_CartesianCoordTo3DPoint.y := #cartesianCoord.y;
   #LKinCtrl_CartesianCoordTo3DPoint.z := #cartesianCoord.z;
END_FUNCTION

FUNCTION "LKinCtrl_3DPointToCartesianCoord" : "LKinCtrl_typeCartesianPosition"   // FC35066, SCL
TITLE = LKinCtrl_3DPointToCartesianCoord
{ S7_Optimized_Access := 'TRUE' }
AUTHOR : tech.team.motioncontrol@siemens.com
FAMILY : LKinCtrl
VERSION : 1.0
// The function converts data type "LKinCtrl_typeCOff3DPoint" in "LKinCtrl_typeCartesianPosition"
   VAR_INPUT
      point3D : "LKinCtrl_typeCOff3DPoint";   // 3D input point
   END_VAR
   // Ret_Val : Return - Cartesian output coordinate
BEGIN
   //==========================================================================================
   // SIEMENS AG
   // (c)Copyright 2019 All Rights Reserved
   //------------------------------------------------------------------------------------------
   // Library: LCOffset
   // Tested with: S7-1515T-3 PN/DP
   // Engineering: TIA Portal V15
   // Restrictions: ---
   // Requirements: S7-1500T FW 2.5
   // Functionality: The function converts data type "LKinCtrl_typeCOff3DPoint" in "LKinCtrl_typeCartesianPosition"
   // Support: tech.team.motioncontrol@siemens.com
   // Note: Parameter comments are only available in language 'English (United States)'
   //------------------------------------------------------------------------------------------
   // Change log table:
   // Version    Date          Expert in charge    Changes applied
   // 01.00.00   2019-02-14    AW                  created
   //===========================================================================================
   //
   #LKinCtrl_3DPointToCartesianCoord.x := #point3D.x;
   #LKinCtrl_3DPointToCartesianCoord.y := #point3D.y;
   #LKinCtrl_3DPointToCartesianCoord.z := #point3D.z;
END_FUNCTION

FUNCTION "LKinCtrl_CalcVecDistancePathPlane" : Word   // FC35067, SCL
TITLE = LKinCtrl_CalcVecDistancePathPlane
{ S7_Optimized_Access := 'TRUE' }
AUTHOR : tech.team.motioncontrol@siemens.com
FAMILY : LKinCtrl
VERSION : 1.0
// Calculate vector distance with respect to path plane
   VAR_INPUT
      vectorInA : "LKinCtrl_typeCOff3DPoint";   // Vector A
      vectorInB : "LKinCtrl_typeCOff3DPoint";   // vector B
      pathPlane : Int;   // Path plane: XZ= 0, YZ=1, XY= 2
   END_VAR
   VAR_OUTPUT
      distancePathPlane : LReal;   // Distance with respect to path plane
   END_VAR
   VAR_TEMP
      tempVectorA : "LKinCtrl_typeCOff3DPoint";
      tempVectorB : "LKinCtrl_typeCOff3DPoint";
   END_VAR
   // Ret_Val : Return value
   VAR CONSTANT
      ERR_COFF_INVALID_PATH_PLANE : Word := 16#8303;   // Error - invalid path plane
   END_VAR
BEGIN
   //=============================================================================
   // SIEMENS AG
   // (c)Copyright 2019 All Rights Reserved
   //-----------------------------------------------------------------------------
   // Library: - 
   // Tested with: S7-1516T-3 PN
   // Engineering: TIA Portal V15
   // Restrictions: -
   // Requirements: S7-1500/S7-1500T FW 2.5
   // Functionality: Calculate vector distance with respect to path plane
   //-----------------------------------------------------------------------------
   // Change log table:
   // Version  Date       Expert in charge Changes applied
   // 01.00.00 2019-02-15 AW               created
   //=============================================================================
   REGION PLAUSIBILITY_CHECK
     // Check path plane
     IF ((#pathPlane >= "CP_XZ") AND (#pathPlane <= "CP_XY"))
     THEN
       ;
     ELSE
       #LKinCtrl_CalcVecDistancePathPlane := #ERR_COFF_INVALID_PATH_PLANE; // Invalid path plane
       RETURN;
     END_IF;
   END_REGION PLAUSIBILITY_CHECK


   REGION CALCULATION
     #tempVectorA := #vectorInA;
     #tempVectorB := #vectorInB;